// TIA Portal project "ROLLINGMILLPLC" (V16) (continued)
VERSION : 0.1
// This block is AUTO GENERATED - DO NOT MODIFY this block!
// Created by Target 1500S version 0
// at 0 
// ********************************************************
//  This is generated by Target 1500S for Simulink
//  Model name:                  LQ
//  Model version:               1.16
//                
//  ODK 1500S version:           V2.5
//  Target 1500S version:        V4.0         
//  MATLAB version:              9.9 (R2020b) 29-Jul-2020
//  Simulink version:            10.2 (R2020b) 29-Jul-2020
//  MATLAB Coder version:        5.1 (R2020b) 29-Jul-2020
//  Simulink Coder version:      9.4 (R2020b) 29-Jul-2020
// 
//  ***Model details***
//  Step Size:                   0.01
//  Default parameter behaviour: Tunable 
//  External Mode:               Off
//  ***ODK 1500S details***  
//  Heap Size:                   32k
//  Max Block Size:              1024
//  Size of thread stack:        32k
//  SyncCallParallelCount:       1(max. number of parallel calls into this ODK application)
//  ********************************************************
// Call this FB to establish a connection to user defined Web page.
   VAR_INPUT
      InternalSignals : "LQInternalModelSignals";
      CTRL_DB : DB_WWW;
   END_VAR
   VAR_IN_OUT
      Params : "LQParams";
   END_VAR
   VAR
      TestPointedSignals : "LQInternalModelSignals";
      Parameter : "LQParams";
      RWParams_Instance : "LQReadWriteParameters";
      Write : Int := 0;
      RunTime : LReal;
   END_VAR
   VAR_TEMP
      ret : Int;
   END_VAR
BEGIN
   // This is generated by Target 1500S for Simulink
   // Model name:                  LQ
   // Model version:               1.16
   //               
   // ODK 1500S version:           V2.5
   // Target 1500S version:        V4.0         
   // MATLAB version:              9.9 (R2020b) 29-Jul-2020
   // Simulink version:            10.2 (R2020b) 29-Jul-2020
   // MATLAB Coder version:        5.1 (R2020b) 29-Jul-2020
   // Simulink Coder version:      9.4 (R2020b) 29-Jul-2020
   //
   // ***Model details***
   // Step Size:                   0.01
   // Default parameter behaviour: Tunable 
   // External Mode:               Off
   // ***ODK 1500S details***  
   // Heap Size:                   32k
   // Max Block Size:              1024
   // Size of thread stack:        32k
   // SyncCallParallelCount:       1(max. number of parallel calls into this ODK application)
   // ********************************************************
   //Call this FB to establish a connection to user defined Web page.
   #RunTime := #RunTime + 10.0;

   #TestPointedSignals := #InternalSignals;
   CASE #Write OF
       0:
           #RWParams_Instance(write := FALSE,
                              STATUS => #RWParams_Instance.STATUS,
                              inOutParams := #Parameter);
           #Params := #Parameter;
       1:
           // Wait for parameter be updated by the Web action
           ;
       2:
           #RWParams_Instance(write := TRUE,
                              STATUS => #RWParams_Instance.STATUS,
                              inOutParams := #Parameter);
           #Params := #Parameter;
           #Write := 0;
       ELSE
           // Not possible to reach
           ;
   END_CASE;

   #ret := WWW(#CTRL_DB);
END_FUNCTION_BLOCK

ORGANIZATION_BLOCK "Main"   // OB1, LAD, ProgramCycle
TITLE = "Main Program Sweep (Cycle)"
{ S7_Optimized_Access := 'TRUE' }
VERSION : 0.1
   VAR_INPUT
      Initial_Call : Bool;   // Initial call of this OB
      Remanence : Bool;   // =True, if remanent data are available
   END_VAR
BEGIN
END_ORGANIZATION_BLOCK

ORGANIZATION_BLOCK "Cyclic interrupt"   // OB30, LAD, CyclicInterrupt
{ S7_Optimized_Access := 'TRUE' }
VERSION : 0.1
   VAR_INPUT
      Initial_Call : Bool;   // Initial call of this OB
      Event_Count : Int;   // Events discarded
   END_VAR
BEGIN

REGION Network 1 (SCL)
   "LQ_GlobalData".Feedback := "OpcInterface".Feedback;
END_REGION

REGION Network 2
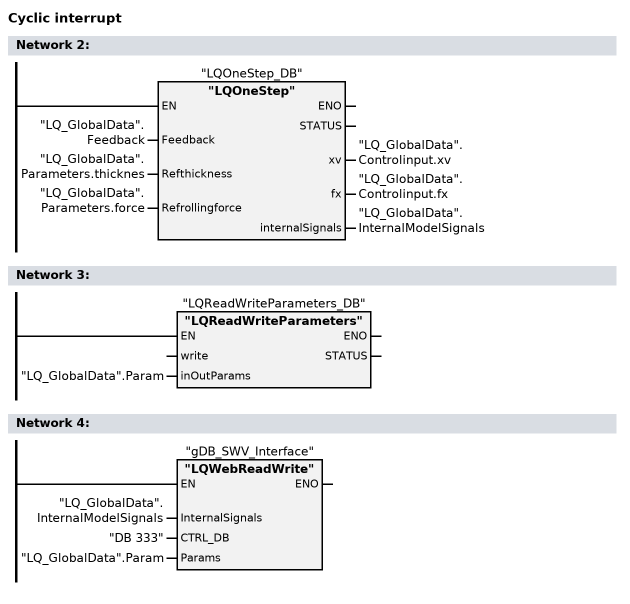
   RUNG wire#powerrail
      "LQOneStep_DB"(Feedback := "LQ_GlobalData".Feedback, Refthickness := "LQ_GlobalData".Parameters.thicknes, Refrollingforce := "LQ_GlobalData".Parameters.force, STATUS =>, xv => "LQ_GlobalData".Controlinput.xv, fx => "LQ_GlobalData".Controlinput.fx, internalSignals => "LQ_GlobalData".InternalModelSignals)
   END_RUNG
   // the same network as SCL:
   "LQOneStep_DB"(Feedback := "LQ_GlobalData".Feedback,   // "LQOneStep"
                  Refthickness := "LQ_GlobalData".Parameters.thicknes,
                  Refrollingforce := "LQ_GlobalData".Parameters.force,
                  xv => "LQ_GlobalData".Controlinput.xv,
                  fx => "LQ_GlobalData".Controlinput.fx,
                  internalSignals => "LQ_GlobalData".InternalModelSignals);
END_REGION

REGION Network 3
   RUNG wire#powerrail
      "LQReadWriteParameters_DB"(write :=, inOutParams := "LQ_GlobalData".Param, STATUS =>)
   END_RUNG
   // the same network as SCL:
   "LQReadWriteParameters_DB"(inOutParams := "LQ_GlobalData".Param);   // "LQReadWriteParameters"
END_REGION

REGION Network 4
   RUNG wire#powerrail
      "gDB_SWV_Interface"(InternalSignals := "LQ_GlobalData".InternalModelSignals, CTRL_DB := "DB 333", Params := "LQ_GlobalData".Param)
   END_RUNG
   // the same network as SCL:
   "gDB_SWV_Interface"(InternalSignals := "LQ_GlobalData".InternalModelSignals,   // "LQWebReadWrite"
                       CTRL_DB := "DB 333",
                       Params := "LQ_GlobalData".Param);
END_REGION

REGION Network 5 (SCL)
   "OpcInterface".Controlinput.xv := "LQ_GlobalData".Controlinput.xv;
   "OpcInterface".Controlinput.fx := "LQ_GlobalData".Controlinput.fx;
END_REGION
END_ORGANIZATION_BLOCK

ORGANIZATION_BLOCK "Startup"   // OB100, LAD, Startup
TITLE = "Complete Restart"
{ S7_Optimized_Access := 'TRUE' }
VERSION : 0.1
   VAR_INPUT
      LostRetentive : Bool;   // True if retentive data are lost
      LostRTC : Bool;   // True if date and time are lost
   END_VAR
BEGIN

REGION Network 1
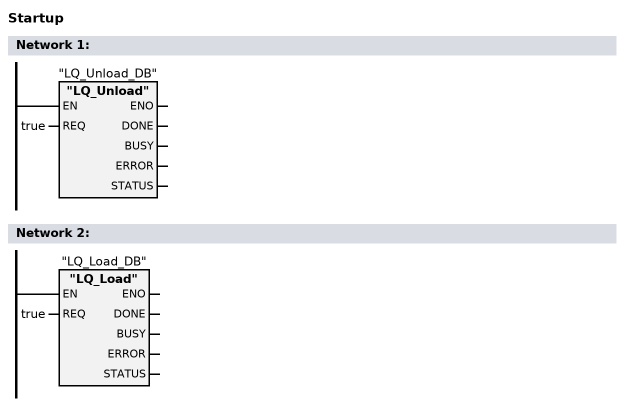
   RUNG wire#powerrail
      "LQ_Unload_DB"(REQ := true, DONE =>, BUSY =>, ERROR =>, STATUS =>)
   END_RUNG
   // the same network as SCL:
   "LQ_Unload_DB"(REQ := true);   // "LQ_Unload"
END_REGION

REGION Network 2
   RUNG wire#powerrail
      "LQ_Load_DB"(REQ := true, DONE =>, BUSY =>, ERROR =>, STATUS =>)
   END_RUNG
   // the same network as SCL:
   "LQ_Load_DB"(REQ := true);   // "LQ_Load"
END_REGION
END_ORGANIZATION_BLOCK

// ===== PLC "PLC_3"  CPU 1518-4 PN/DP MFP =====

TYPE "LQInternalModelSignals"
// This block is AUTO GENERATED - DO NOT MODIFY this block!
// Created by ODK_CodeGenerator version 205.100.101.18
// at Fri August 27 01:33:44 2021
// ********************************************************
   STRUCT
      Controlinput : Array[0..1] of LReal;
      Feedback : Array[0..4] of LReal;
      LQ_Refthickness : LReal;
      LQ_Refrollingforce : LReal;
   END_STRUCT;
END_TYPE

TYPE "LQParams"
// This block is AUTO GENERATED - DO NOT MODIFY this block!
// Created by ODK_CodeGenerator version 205.100.101.18
// at Mon August 30 17:02:50 2021
// ********************************************************
   STRUCT
      Lr : Array[0..3] of LReal;   // [LQ Controller 1/Gain Lr]:LQ_P.Lr
      Ly : Array[0..9] of LReal;   // [LQ Controller 1/Gain Ly]:LQ_P.Ly
   END_STRUCT;
   // Lr[0] := 0.013106;
   // Lr[1] := 0.0;
   // Lr[2] := 0.0;
   // Lr[3] := 3.112673;
   // Ly[0] := 0.0;
   // Ly[1] := 0.0;
   // Ly[2] := 0.0;
   // Ly[3] := 0.0;
   // Ly[4] := 0.011684;
   // Ly[5] := 0.0;
   // Ly[6] := 3.8E-05;
   // Ly[7] := 0.0;
   // Ly[8] := 0.0;
   // Ly[9] := 3.112673;
END_TYPE

DATA_BLOCK "LQ_GlobalData"   // DB1
{ S7_Optimized_Access := 'TRUE' }
VERSION : 0.1
   VAR
      Parameters : Struct
         thicknes : LReal;
         force : LReal;
      END_STRUCT;
      Feedback : Array[0..4] of LReal;
      Controlinput : Struct
         xv : LReal;
         fx : LReal;
      END_STRUCT;
      InternalModelSignals : "LQInternalModelSignals";
   END_VAR
   VAR RETAIN
      Param : "LQParams";
   END_VAR
BEGIN
END_DATA_BLOCK

DATA_BLOCK "gDB_SWV_Interface"   // DB2
{ S7_Optimized_Access := 'TRUE' }
VERSION : 0.1
// stored: InstanceOfName LQWebReadWrite
"LQWebReadWrite"
BEGIN
END_DATA_BLOCK

DATA_BLOCK "OpcInterface"   // DB3
{ S7_Optimized_Access := 'TRUE' }
VERSION : 0.1
   VAR
      Feedback : Array[0..4] of LReal;
      Controlinput : Struct
         xv : LReal;
         fx : LReal;
      END_STRUCT;
   END_VAR
BEGIN
END_DATA_BLOCK

DATA_BLOCK "LQ_Load_DB"   // DB4
{ S7_Optimized_Access := 'TRUE' }
VERSION : 0.1
// stored: InstanceOfName LQ_Load
"LQ_Load"
BEGIN
END_DATA_BLOCK

DATA_BLOCK "LQOneStep_DB"   // DB5
{ S7_Optimized_Access := 'TRUE' }
VERSION : 0.1
// stored: InstanceOfName LQOneStep
"LQOneStep"
BEGIN
END_DATA_BLOCK

DATA_BLOCK "LQReadWriteParameters_DB"   // DB6
{ S7_Optimized_Access := 'TRUE' }
VERSION : 0.1
// stored: InstanceOfName LQReadWriteParameters
"LQReadWriteParameters"
BEGIN
END_DATA_BLOCK

DATA_BLOCK "LQ_Unload_DB"   // DB7
{ S7_Optimized_Access := 'TRUE' }
VERSION : 0.1
// stored: InstanceOfName LQ_Unload
"LQ_Unload"
BEGIN
END_DATA_BLOCK

FUNCTION_BLOCK "LQ_Load"   // FB1, SCL
{ S7_Optimized_Access := 'TRUE' }
VERSION : 0.1
// This block is AUTO GENERATED - DO NOT MODIFY this block!
// Created by ODK_CodeGenerator version 2.5.1
// at Fri August 27 01:33:44 2021
// max. number of parallel calls into this ODK application is: 1
// *************************************************************
   VAR_INPUT
      REQ : Bool;
   END_VAR
   VAR_OUTPUT
      DONE : Bool;
      BUSY : Bool;
      ERROR : Bool;
      STATUS : Int;
   END_VAR
   VAR
      ODK_Load_Instance : ODK_Load;
      _odk_internal_LIBRARY_NAME : String := '<rt>LQ_ODK.so';
   END_VAR
   VAR CONSTANT
      _odk_internal_INSTANCE_ID : UDInt := 101_277_234;
   END_VAR
BEGIN
   //
   // DO NOT CHANGE BELOW OF THIS LINE !!
   // This is an automatic generated block by the
   // SIMATIC ODK 1500S V2.5.1
   // DO NOT CHANGE !!
   //
   #ODK_Load_Instance(REQ := #REQ,
                      LIBRARY_NAME := #_odk_internal_LIBRARY_NAME,
                      INSTANCE_ID := #_odk_internal_INSTANCE_ID,
                      DONE => #DONE,
                      BUSY => #BUSY,
                      ERROR => #ERROR,
                      STATUS => #STATUS);
   //
   // DO NOT CHANGE !!
   // This is an automatic generated block by the
   // SIMATIC ODK 1500S V2.5.1
   // DO NOT CHANGE ABOVE OF THIS LINE !!
   //
END_FUNCTION_BLOCK

FUNCTION_BLOCK "LQ_Unload"   // FB2, SCL
{ S7_Optimized_Access := 'TRUE' }
VERSION : 0.1
// This block is AUTO GENERATED - DO NOT MODIFY this block!
// Created by ODK_CodeGenerator version 205.100.101.18
// at Fri August 27 01:33:44 2021
// max. number of parallel calls into this ODK application is: 1
// *************************************************************
   VAR_INPUT
      REQ : Bool;
   END_VAR
   VAR_OUTPUT
      DONE : Bool;
      BUSY : Bool;
      ERROR : Bool;
      STATUS : Int;
   END_VAR
   VAR
      ODK_Unld_Instance : ODK_Unld;
   END_VAR
   VAR CONSTANT
      _odk_internal_INSTANCE_ID : UDInt := 101_277_234;
   END_VAR
BEGIN
   //
   // DO NOT CHANGE BELOW OF THIS LINE !!
   // This is an automatic generated block by the
   // SIMATIC ODK 1500S V2.5.1
   // DO NOT CHANGE !!
   //
   #ODK_Unld_Instance(REQ := #REQ,
                      INSTANCE_ID := #_odk_internal_INSTANCE_ID,
                      DONE => #DONE,
                      BUSY => #BUSY,
                      ERROR => #ERROR,
                      STATUS => #STATUS);
   //
   // DO NOT CHANGE !!
   // This is an automatic generated block by the
   // SIMATIC ODK 1500S V2.5.1
   // DO NOT CHANGE ABOVE OF THIS LINE !!
   //
END_FUNCTION_BLOCK

FUNCTION_BLOCK "LQOneStep"   // FB3, SCL
{ S7_Optimized_Access := 'TRUE' }
VERSION : 0.1
// This block is AUTO GENERATED - DO NOT MODIFY this block!
// Created by ODK_CodeGenerator version 205.100.101.18
// at Fri August 27 01:33:44 2021
// max. number of parallel calls into this ODK application is: 1
// *************************************************************
//  This is generated by Target 1500S for Simulink
//  Model name:                  LQ
//  Model version:               1.16
//                 
//  ODK 1500S version:           V2.5
//  Target 1500S version:        V4.0         
//  MATLAB version:              9.9 (R2020b) 29-Jul-2020
//  Simulink version:            10.2 (R2020b) 29-Jul-2020
//  MATLAB Coder version:        5.1 (R2020b) 29-Jul-2020
//  Simulink Coder version:      9.4 (R2020b) 29-Jul-2020
//  
//  ***Model details***
//  Step Size:                   0.01
//  Default parameter behaviour: Tunable
//  External Mode:               Off
//  
//  ***ODK 1500S details***  
//  Heap Size:                   32k
//  Max Block Size:              1024
//  Size of thread stack:        32k
//  SyncCallParallelCount:       1(max. number of parallel calls into this ODK application)
//  ********************************************************
   VAR_INPUT
      Feedback : Array[0..4] of LReal;
      Refthickness : LReal;
      Refrollingforce : LReal;
   END_VAR
   VAR_OUTPUT
      STATUS : Int := 0;
      xv : LReal;
      fx : LReal;
      internalSignals : "LQInternalModelSignals";
   END_VAR
   VAR
      _odk_internal_Last_REQ : Bool := FALSE;
      _odk_internal_Last_BUSY : Bool := FALSE;
      _odk_internal_IN_BUFFER : Array[0..55] of Byte;
      _odk_internal_OUT_BUFFER : Array[0..87] of Byte;
   END_VAR
   VAR_TEMP
      _odk_internal_pos : DInt;
      _odk_internal_err : Int;
      _odk_internal_i : Int;
   END_VAR
   VAR CONSTANT
      _odk_internal_INSTANCE_ID : UDInt := 101_277_234;
      _odk_internal_COMMAND : UDInt := 295_977_560;
   END_VAR
BEGIN
   //
   // DO NOT CHANGE BELOW OF THIS LINE !!
   // This is an automatic generated block by the
   // SIMATIC ODK 1500S V2.5.1
   // DO NOT CHANGE !!
   //
   // This is generated by Target 1500S for Simulink
   // Model name:                  LQ
   // Model version:               1.16
   //                
   // ODK 1500S version:           V2.5
   // Target 1500S version:        V4.0         
   // MATLAB version:              9.9 (R2020b) 29-Jul-2020
   // Simulink version:            10.2 (R2020b) 29-Jul-2020
   // MATLAB Coder version:        5.1 (R2020b) 29-Jul-2020
   // Simulink Coder version:      9.4 (R2020b) 29-Jul-2020
   // 
   // ***Model details***
   // Step Size:                   0.01
   // Default parameter behaviour: Tunable
   // External Mode:               Off
   // 
   // ***ODK 1500S details***  
   // Heap Size:                   32k
   // Max Block Size:              1024
   // Size of thread stack:        32k
   // SyncCallParallelCount:       1(max. number of parallel calls into this ODK application)
   // ********************************************************
   // 
   #_odk_internal_pos := 0;
   FOR #_odk_internal_i := 0 TO 4 DO
       #_odk_internal_err := WRITE_LITTLE(src_variable := #Feedback[#_odk_internal_i], dest_array := #_odk_internal_IN_BUFFER, pos := #_odk_internal_pos);
   END_FOR;
   #_odk_internal_err := WRITE_LITTLE(src_variable := #Refthickness, dest_array := #_odk_internal_IN_BUFFER, pos := #_odk_internal_pos);
   #_odk_internal_err := WRITE_LITTLE(src_variable := #Refrollingforce, dest_array := #_odk_internal_IN_BUFFER, pos := #_odk_internal_pos);
   #STATUS := ODK_ExcS(INSTANCE_ID := #_odk_internal_INSTANCE_ID,
                       COMMAND := #_odk_internal_COMMAND,
                       IN_DATA := #_odk_internal_IN_BUFFER,
                       INOUT_DATA := null,
                       OUT_DATA := #_odk_internal_OUT_BUFFER
   );
   IF INT_TO_UINT(#STATUS) < 16#7000 THEN
       #_odk_internal_pos := 0;
       #_odk_internal_err := READ_LITTLE(dest_Variable => #xv, src_array := #_odk_internal_OUT_BUFFER, pos := #_odk_internal_pos);
       #_odk_internal_err := READ_LITTLE(dest_Variable => #fx, src_array := #_odk_internal_OUT_BUFFER, pos := #_odk_internal_pos);
       FOR #_odk_internal_i := 0 TO 1 DO
           #_odk_internal_err := READ_LITTLE(dest_Variable => #internalSignals.#Controlinput[#_odk_internal_i], src_array := #_odk_internal_OUT_BUFFER, pos := #_odk_internal_pos);
       END_FOR;
       FOR #_odk_internal_i := 0 TO 4 DO
           #_odk_internal_err := READ_LITTLE(dest_Variable => #internalSignals.#Feedback[#_odk_internal_i], src_array := #_odk_internal_OUT_BUFFER, pos := #_odk_internal_pos);
       END_FOR;
       #_odk_internal_err := READ_LITTLE(dest_Variable => #internalSignals.#LQ_Refthickness, src_array := #_odk_internal_OUT_BUFFER, pos := #_odk_internal_pos);
       #_odk_internal_err := READ_LITTLE(dest_Variable => #internalSignals.#LQ_Refrollingforce, src_array := #_odk_internal_OUT_BUFFER, pos := #_odk_internal_pos);
   END_IF;
   //
   // DO NOT CHANGE !!
   // This is an automatic generated block by the
   // SIMATIC ODK 1500S V2.5.1
   // DO NOT CHANGE ABOVE OF THIS LINE !!
   //
END_FUNCTION_BLOCK

FUNCTION_BLOCK "LQReadWriteParameters"   // FB4, SCL
{ S7_Optimized_Access := 'TRUE' }
VERSION : 0.1
// This block is AUTO GENERATED - DO NOT MODIFY this block!
// Created by ODK_CodeGenerator version 205.100.101.18
// at Fri August 27 01:33:44 2021
// max. number of parallel calls into this ODK application is: 1
// *************************************************************
//  This is generated by Target 1500S for Simulink
//  Model name:                  LQ
//  Model version:               1.16
//                 
//  ODK 1500S version:           V2.5
//  Target 1500S version:        V4.0         
//  MATLAB version:              9.9 (R2020b) 29-Jul-2020
//  Simulink version:            10.2 (R2020b) 29-Jul-2020
//  MATLAB Coder version:        5.1 (R2020b) 29-Jul-2020
//  Simulink Coder version:      9.4 (R2020b) 29-Jul-2020
//  
//  ***Model details***
//  Step Size:                   0.01
//  Default parameter behaviour: Tunable
//  External Mode:               Off
//  
//  ***ODK 1500S details***  
//  Heap Size:                   32k
//  Max Block Size:              1024
//  Size of thread stack:        32k
//  SyncCallParallelCount:       1(max. number of parallel calls into this ODK application)
//  ********************************************************
//  
//  Call this function to read or write parameters from/to Simulink Model.
//  Set write[IN] parameter to TRUE in order to write and set FALSE to read parameters
   VAR_INPUT
      write : Bool;
   END_VAR
   VAR_OUTPUT
      STATUS : Int := 0;
   END_VAR
   VAR_IN_OUT
      inOutParams : "LQParams";
   END_VAR
   VAR
      _odk_internal_Last_REQ : Bool := FALSE;
      _odk_internal_Last_BUSY : Bool := FALSE;
      _odk_internal_IN_BUFFER : Array[0..0] of Byte;
      _odk_internal_INOUT_BUFFER : Array[0..111] of Byte;
   END_VAR
   VAR_TEMP
      _odk_internal_pos : DInt;
      _odk_internal_err : Int;
      _odk_internal_i : Int;
   END_VAR
   VAR CONSTANT
      _odk_internal_INSTANCE_ID : UDInt := 101_277_234;
      _odk_internal_COMMAND : UDInt := 2_137_970_399;
   END_VAR
BEGIN
   //
   // DO NOT CHANGE BELOW OF THIS LINE !!
   // This is an automatic generated block by the
   // SIMATIC ODK 1500S V2.5.1
   // DO NOT CHANGE !!
   //
   // This is generated by Target 1500S for Simulink
   // Model name:                  LQ
   // Model version:               1.16
   //                
   // ODK 1500S version:           V2.5
   // Target 1500S version:        V4.0         
   // MATLAB version:              9.9 (R2020b) 29-Jul-2020
   // Simulink version:            10.2 (R2020b) 29-Jul-2020
   // MATLAB Coder version:        5.1 (R2020b) 29-Jul-2020
   // Simulink Coder version:      9.4 (R2020b) 29-Jul-2020
   // 
   // ***Model details***
   // Step Size:                   0.01
   // Default parameter behaviour: Tunable
   // External Mode:               Off
   // 
   // ***ODK 1500S details***  
   // Heap Size:                   32k
   // Max Block Size:              1024
   // Size of thread stack:        32k
   // SyncCallParallelCount:       1(max. number of parallel calls into this ODK application)
   // ********************************************************
   // 
   // Call this function to read or write parameters from/to Simulink Model.
   // Set write[IN] parameter to TRUE in order to write and set FALSE to read parameters
   #_odk_internal_pos := 0;
   IF (True = #write) THEN
       #_odk_internal_IN_BUFFER[#_odk_internal_pos] := BYTE#1;
   ELSE
       #_odk_internal_IN_BUFFER[#_odk_internal_pos] := BYTE#0;
   END_IF;
   #_odk_internal_pos := #_odk_internal_pos + 1;
   #_odk_internal_pos := 0;
   FOR #_odk_internal_i := 0 TO 3 DO
       #_odk_internal_err := WRITE_LITTLE(src_variable := #inOutParams.#Lr[#_odk_internal_i], dest_array := #_odk_internal_INOUT_BUFFER, pos := #_odk_internal_pos);
   END_FOR;
   FOR #_odk_internal_i := 0 TO 9 DO
       #_odk_internal_err := WRITE_LITTLE(src_variable := #inOutParams.#Ly[#_odk_internal_i], dest_array := #_odk_internal_INOUT_BUFFER, pos := #_odk_internal_pos);
   END_FOR;
   #STATUS := ODK_ExcS(INSTANCE_ID := #_odk_internal_INSTANCE_ID,
                       COMMAND := #_odk_internal_COMMAND,
                       IN_DATA := #_odk_internal_IN_BUFFER,
                       INOUT_DATA := #_odk_internal_INOUT_BUFFER,
                       OUT_DATA := null);
   IF INT_TO_UINT(#STATUS) < 16#7000 THEN
       #_odk_internal_pos := 0;
       FOR #_odk_internal_i := 0 TO 3 DO
           #_odk_internal_err := READ_LITTLE(dest_Variable => #inOutParams.#Lr[#_odk_internal_i], src_array := #_odk_internal_INOUT_BUFFER, pos := #_odk_internal_pos);
       END_FOR;
       FOR #_odk_internal_i := 0 TO 9 DO
           #_odk_internal_err := READ_LITTLE(dest_Variable => #inOutParams.#Ly[#_odk_internal_i], src_array := #_odk_internal_INOUT_BUFFER, pos := #_odk_internal_pos);
       END_FOR;
   END_IF;
   //
   // DO NOT CHANGE !!
   // This is an automatic generated block by the
   // SIMATIC ODK 1500S V2.5.1
   // DO NOT CHANGE ABOVE OF THIS LINE !!
   //
END_FUNCTION_BLOCK

FUNCTION_BLOCK "LQWebReadWrite"   // FB5, SCL
{ S7_Optimized_Access := 'TRUE' }
VERSION : 0.1
// This block is AUTO GENERATED - DO NOT MODIFY this block!
// Created by Target 1500S version 0
// at 0 
// ********************************************************
//  This is generated by Target 1500S for Simulink
//  Model name:                  LQ
//  Model version:               1.16
//                
//  ODK 1500S version:           V2.5
//  Target 1500S version:        V4.0         
//  MATLAB version:              9.9 (R2020b) 29-Jul-2020
//  Simulink version:            10.2 (R2020b) 29-Jul-2020
//  MATLAB Coder version:        5.1 (R2020b) 29-Jul-2020
//  Simulink Coder version:      9.4 (R2020b) 29-Jul-2020
// 
//  ***Model details***
//  Step Size:                   0.01
//  Default parameter behaviour: Tunable 
//  External Mode:               Off
//  ***ODK 1500S details***  
//  Heap Size:                   32k
//  Max Block Size:              1024
//  Size of thread stack:        32k
//  SyncCallParallelCount:       1(max. number of parallel calls into this ODK application)
//  ********************************************************
// Call this FB to establish a connection to user defined Web page.
   VAR_INPUT
      InternalSignals : "LQInternalModelSignals";
      CTRL_DB : DB_WWW;
   END_VAR
   VAR_IN_OUT
      Params : "LQParams";
   END_VAR
   VAR
      TestPointedSignals : "LQInternalModelSignals";
      Parameter : "LQParams";
      RWParams_Instance : "LQReadWriteParameters";
      Write : Int := 0;
      RunTime : LReal;
   END_VAR
   VAR_TEMP
      ret : Int;
   END_VAR
BEGIN
   // This is generated by Target 1500S for Simulink
   // Model name:                  LQ
   // Model version:               1.16
   //               
   // ODK 1500S version:           V2.5
   // Target 1500S version:        V4.0         
   // MATLAB version:              9.9 (R2020b) 29-Jul-2020
   // Simulink version:            10.2 (R2020b) 29-Jul-2020
   // MATLAB Coder version:        5.1 (R2020b) 29-Jul-2020
   // Simulink Coder version:      9.4 (R2020b) 29-Jul-2020
   //
   // ***Model details***
   // Step Size:                   0.01
   // Default parameter behaviour: Tunable 
   // External Mode:               Off
   // ***ODK 1500S details***  
   // Heap Size:                   32k
   // Max Block Size:              1024
   // Size of thread stack:        32k
   // SyncCallParallelCount:       1(max. number of parallel calls into this ODK application)
   // ********************************************************
   //Call this FB to establish a connection to user defined Web page.
   #RunTime := #RunTime + 10.0;

   #TestPointedSignals := #InternalSignals;
   CASE #Write OF
       0:
           #RWParams_Instance(write := FALSE,
                              STATUS => #RWParams_Instance.STATUS,
                              inOutParams := #Parameter);
           #Params := #Parameter;
       1:
           // Wait for parameter be updated by the Web action
           ;
       2:
           #RWParams_Instance(write := TRUE,
                              STATUS => #RWParams_Instance.STATUS,
                              inOutParams := #Parameter);
           #Params := #Parameter;
           #Write := 0;
       ELSE
           // Not possible to reach
           ;
   END_CASE;

   #ret := WWW(#CTRL_DB);
END_FUNCTION_BLOCK

ORGANIZATION_BLOCK "Main"   // OB1, LAD, ProgramCycle
TITLE = "Main Program Sweep (Cycle)"
{ S7_Optimized_Access := 'TRUE' }
VERSION : 0.1
   VAR_INPUT
      Initial_Call : Bool;   // Initial call of this OB
      Remanence : Bool;   // =True, if remanent data are available
   END_VAR
BEGIN
END_ORGANIZATION_BLOCK

ORGANIZATION_BLOCK "Cyclic interrupt"   // OB30, LAD, CyclicInterrupt
{ S7_Optimized_Access := 'TRUE' }
VERSION : 0.1
   VAR_INPUT
      Initial_Call : Bool;   // Initial call of this OB
      Event_Count : Int;   // Events discarded
   END_VAR
BEGIN

REGION Network 1 (SCL)
   "LQ_GlobalData".Feedback := "OpcInterface".Feedback;
END_REGION

REGION Network 2
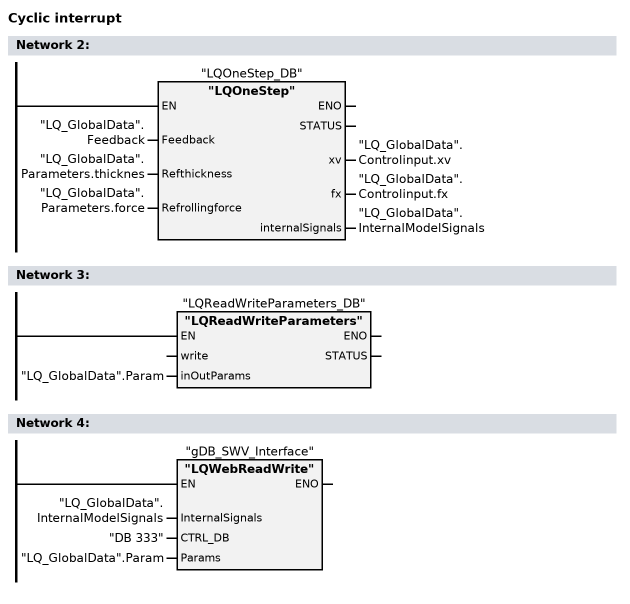
   RUNG wire#powerrail
      "LQOneStep_DB"(Feedback := "LQ_GlobalData".Feedback, Refthickness := "LQ_GlobalData".Parameters.thicknes, Refrollingforce := "LQ_GlobalData".Parameters.force, STATUS =>, xv => "LQ_GlobalData".Controlinput.xv, fx => "LQ_GlobalData".Controlinput.fx, internalSignals => "LQ_GlobalData".InternalModelSignals)
   END_RUNG
   // the same network as SCL:
   "LQOneStep_DB"(Feedback := "LQ_GlobalData".Feedback,   // "LQOneStep"
                  Refthickness := "LQ_GlobalData".Parameters.thicknes,
                  Refrollingforce := "LQ_GlobalData".Parameters.force,
                  xv => "LQ_GlobalData".Controlinput.xv,
                  fx => "LQ_GlobalData".Controlinput.fx,
                  internalSignals => "LQ_GlobalData".InternalModelSignals);
END_REGION

REGION Network 3
   RUNG wire#powerrail
      "LQReadWriteParameters_DB"(write :=, inOutParams := "LQ_GlobalData".Param, STATUS =>)
   END_RUNG
   // the same network as SCL:
   "LQReadWriteParameters_DB"(inOutParams := "LQ_GlobalData".Param);   // "LQReadWriteParameters"
END_REGION

REGION Network 4
   RUNG wire#powerrail
      "gDB_SWV_Interface"(InternalSignals := "LQ_GlobalData".InternalModelSignals, CTRL_DB := "DB 333", Params := "LQ_GlobalData".Param)
   END_RUNG
   // the same network as SCL:
   "gDB_SWV_Interface"(InternalSignals := "LQ_GlobalData".InternalModelSignals,   // "LQWebReadWrite"
                       CTRL_DB := "DB 333",
                       Params := "LQ_GlobalData".Param);
END_REGION

REGION Network 5 (SCL)
   "OpcInterface".Controlinput.xv := "LQ_GlobalData".Controlinput.xv;
   "OpcInterface".Controlinput.fx := "LQ_GlobalData".Controlinput.fx;
END_REGION
END_ORGANIZATION_BLOCK

ORGANIZATION_BLOCK "Startup"   // OB100, LAD, Startup
TITLE = "Complete Restart"
{ S7_Optimized_Access := 'TRUE' }
VERSION : 0.1
   VAR_INPUT
      LostRetentive : Bool;   // True if retentive data are lost
      LostRTC : Bool;   // True if date and time are lost
   END_VAR
BEGIN

REGION Network 1
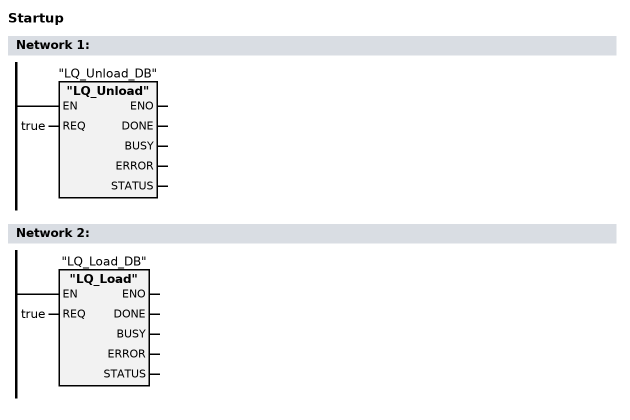
   RUNG wire#powerrail
      "LQ_Unload_DB"(REQ := true, DONE =>, BUSY =>, ERROR =>, STATUS =>)
   END_RUNG
   // the same network as SCL:
   "LQ_Unload_DB"(REQ := true);   // "LQ_Unload"
END_REGION

REGION Network 2
   RUNG wire#powerrail
      "LQ_Load_DB"(REQ := true, DONE =>, BUSY =>, ERROR =>, STATUS =>)
   END_RUNG
   // the same network as SCL:
   "LQ_Load_DB"(REQ := true);   // "LQ_Load"
END_REGION
END_ORGANIZATION_BLOCK

(* ===== HMI "HMI_RT_2" =====
system functions are stored by id; their names below are inferred from use
connection "HMI_Connection_1": ETHERNET, S7_1500_OMS
connection "HMI_Connection_2": ETHERNET, S7_1500_OMS
connection "HMI_Connection_3": ETHERNET, S7_1500_OMS

HMI tags "Default tag table"
   "Tag_ScreenNumber" : UInt, internal
   "LQ_GlobalData_Parameters_thicknes" : LReal = PLC LQ_GlobalData.Parameters.thicknes, 1 s
   "LQ_GlobalData_Parameters_force" : LReal = PLC LQ_GlobalData.Parameters.force, 1 s
   "LQ_GlobalData_Feedback{2}" : LReal = PLC LQ_GlobalData.Feedback[2], 1 s
   "LQ_GlobalData_Parameters_thicknes(1)" : LReal = PLC LQ_GlobalData.Parameters.thicknes, 1 s
   "LQ_GlobalData_Feedback{2}(1)" : LReal = PLC LQ_GlobalData.Feedback[2], 1 s
   "LQ_GlobalData_Parameters_force(1)" : LReal = PLC LQ_GlobalData.Parameters.force, 1 s
   "LQ_GlobalData_Parameters_thicknes(2)" : LReal = PLC LQ_GlobalData.Parameters.thicknes, 1 s
   "LQ_GlobalData_Parameters_force(2)" : LReal = PLC LQ_GlobalData.Parameters.force, 1 s
   "LQ_GlobalData_Feedback{2}(2)" : LReal = PLC LQ_GlobalData.Feedback[2], 1 s
   "LQ_GlobalData_Feedback{4}" : LReal = PLC LQ_GlobalData.Feedback[4], 1 s
   "LQ_GlobalData_Feedback{4}(1)" : LReal = PLC LQ_GlobalData.Feedback[4], 1 s
   "LQ_GlobalData_Feedback{4}(2)" : LReal = PLC LQ_GlobalData.Feedback[4], 1 s

screen "Home" 1280x740, template "Template_1"
   on GenerateScreen: SetTag("Tag_ScreenNumber", 1)
   TextField "HmiScreenItemData_3" at 413,45 size 404x37; Text 'Welcome to HMI of the Rolling Mill'
   Button "HmiScreenItemData" at 471,181 size 159x47; TextOn 'Rolling Stand 1'; TextOff 'Rolling Stand 1'; PictureOn "Navigates to Roller 1 for TP1500 Comfort 16.0.0.0"; PictureOff "Navigates to Roller 1 for TP1500 Comfort 16.0.0.0"
      on Release: ActivateScreen("Rolling Stand 1", 0)
   Button "HmiScreenItemData_1" at 471,261 size 159x47; TextOn 'Rolling Stand 2'; TextOff 'Rolling Stand 2'; PictureOn "Navigates to Roller 2 for TP1500 Comfort 16.0.0.0"; PictureOff "Navigates to Roller 2 for TP1500 Comfort 16.0.0.0"
      on Release: ActivateScreen("Rolling Stand 2", 0)
   Button "HmiScreenItemData_2" at 471,342 size 159x47; TextOn 'Rolling Stand 3'; TextOff 'Rolling Stand 3'; PictureOn "Navigates to Roller 3 for TP1500 Comfort 16.0.0.0"; PictureOff "Navigates to Roller 3 for TP1500 Comfort 16.0.0.0"
      on Release: ActivateScreen("Rolling Stand 3", 0)
   Button "HmiScreenItemData_4" at 538,476 size 159x47; TextOn 'System screens'; TextOff 'System screens'; PictureOn "Navigates to System screens for TP1500 Comfort 16.0.0.0"; PictureOff "Navigates to System screens for TP1500 Comfort 16.0.0.0"
      on Release: ActivateScreen("System screens", 0)
   TextField "Text field_1" at 482,193 size 30x18; Text 'R-1'
   TextField "Text field_2" at 482,275 size 30x18; Text 'R-2'
   TextField "Text field_3" at 482,356 size 30x18; Text 'R-3'
   TextField "Text field_5" at 553,432 size 135x25; Text 'Information'
   Switch "Switch_1" at 683,171 size 77x50; CaptionText 'Switch'; TextOff 'OFF'; TextOn 'ON'
      on SwitchOn: function_f249594b("HMI_Connection_1", 8)
      on SwitchOff: function_f249594b("HMI_Connection_1", 4)
   Switch "Switch_2" at 683,255 size 77x50; TextOn 'ON'; CaptionText 'Switch'; TextOff 'OFF'
      on SwitchOn: function_f249594b("HMI_Connection_2", 8)
      on SwitchOff: function_f249594b("HMI_Connection_2", 4)
   Switch "Switch_3" at 683,335 size 77x50; TextOn 'ON'; CaptionText 'Switch'; TextOff 'OFF'
      on SwitchOn: function_f249594b("HMI_Connection_3", 8)
      on SwitchOff: function_f249594b("HMI_Connection_3", 4)
   TextField "Text field_4" at 480,132 size 110x25; Text 'Mill Stands'
   TextField "Text field_6" at 675,132 size 92x25; Text 'PLC Switch'

screen "Rolling Stand 1" 1280x740, template "Template_1"
   on GenerateScreen: SetTag("Tag_ScreenNumber", 2)
   TextField "HmiScreenItemData" at 146,334 size 1024x27; Text 'Roller 1'
   Button "Back" at 1,25 size 159x47; TextOn 'Back'; TextOff 'Back'
      on Release: ActivateScreen("Home", 0)
   TrendView "Trend view_1" at 295,23 size 984x343
   TextField "Text field_4" at 41,188 size 164x40; Text 'Enter Setpoint'
   Group "Group" at 29,242 size 182x37; FormatPattern 9
   Group "Group_1" at 26,92 size 196x56
   IOField "I/O field_2" at 162,288 size 71x37; FormatPattern 999; Unit N
      ProcessValue <- "LQ_GlobalData_Parameters_force"
   TextField "Text field_3" at 25,288 size 137x37; Text 'Rolling force :'
   TrendView "Trend view_2" at 296,361 size 984x320
   IOField "I/O field_1" at 150,242 size 61x37; FormatPattern 9; Unit mm
      ProcessValue <- "LQ_GlobalData_Parameters_thicknes"
   TextField "Text field_1" at 29,242 size 121x37; Text 'Thickness :'
   TextField "Text field_2" at 26,94 size 196x53; Text 'Rolling Stand 1'

screen "System screens" 1280x740, template "Template_1"
   on GenerateScreen: SetTag("Tag_ScreenNumber", 5)
   Button "Back" at 1,25 size 159x47; TextOn 'Back'; TextOff 'Back'
      on Release: ActivateScreen("Home", 0)
   Button "HmiScreenItemData" at 36,119 size 159x47; TextOn 'SIMATIC PLC system diagnos...'; TextOff 'SIMATIC PLC system diagnos...'; PictureOn "Navigates to SIMATIC PLC system diagnostics for TP1500 Comfort 16.0.0.0"; PictureOff "Navigates to SIMATIC PLC system diagnostics for TP1500 Comfort 16.0.0.0"
      on Release: ActivateScreen("SIMATIC PLC system diagnostics", 0)
   Button "HmiScreenItemData_1" at 36,178 size 159x47; TextOn 'Project information'; TextOff 'Project information'; PictureOn "Navigates to Project information for TP1500 Comfort 16.0.0.0"; PictureOff "Navigates to Project information for TP1500 Comfort 16.0.0.0"
      on Release: ActivateScreen("Project information", 0)
   Button "HmiScreenItemData_2" at 36,237 size 159x47; TextOn 'System settings'; TextOff 'System settings'; PictureOn "Navigates to System settings for TP1500 Comfort 16.0.0.0"; PictureOff "Navigates to System settings for TP1500 Comfort 16.0.0.0"
      on Release: ActivateScreen("System settings", 0)
   Button "HmiScreenItemData_3" at 36,296 size 159x47; TextOn 'User administration'; TextOff 'User administration'; PictureOn "Navigates to User administration for TP1500 Comfort 16.0.0.0"; PictureOff "Navigates to User administration for TP1500 Comfort 16.0.0.0"
      on Release: ActivateScreen("User administration", 0)
   Button "HmiScreenItemData_4" at 36,355 size 159x47; TextOn 'System information'; TextOff 'System information'; PictureOn "Navigates to System information for TP1500 Comfort 16.0.0.0"; PictureOff "Navigates to System information for TP1500 Comfort 16.0.0.0"
      on Release: ActivateScreen("System information", 0)
   Button "HmiScreenItemData_5" at 36,414 size 159x47; TextOn 'Different jobs'; TextOff 'Different jobs'; PictureOn "Navigates to Different jobs for TP1500 Comfort 16.0.0.0"; PictureOff "Navigates to Different jobs for TP1500 Comfort 16.0.0.0"
      on Release: ActivateScreen("Different jobs", 0)

screen "SIMATIC PLC system diagnostics" 1280x740, template "Template_1"
   on GenerateScreen: SetTag("Tag_ScreenNumber", 6)
   SysDiagControl "HmiScreenItemData" at 1,73 size 1276x599
   Button "Back" at 1,25 size 159x47; TextOn 'Back'; TextOff 'Back'
      on Release: ActivateScreen("System screens", 0)

screen "Project information" 1280x740, template "Template_1"
   on GenerateScreen: SetTag("Tag_ScreenNumber", 7)
   TextField "HmiScreenItemData" at 35,75 size 171x28; Text 'Project name:'
   TextField "HmiScreenItemData_1" at 241,75 size 1004x28; Text 'Rolling_Mill_With_Three_Rollers'
   TextField "HmiScreenItemData_2" at 35,105 size 171x28; Text 'Created on:'
   TextField "HmiScreenItemData_3" at 241,105 size 1004x28; Text '5/28/2021 9:23:35 PM'
   TextField "HmiScreenItemData_4" at 35,135 size 171x28; Text 'Author:'
   TextField "HmiScreenItemData_5" at 241,135 size 1004x28; Text 'Mehrab'
   TextField "HmiScreenItemData_6" at 35,165 size 171x28; Text 'Description:'
   TextField "HmiScreenItemData_7" at 241,165 size 1004x28; Text '(not configured)'
   Button "Back" at 1,25 size 159x47; TextOn 'Back'; TextOff 'Back'
      on Release: ActivateScreen("System screens", 0)

screen "System settings" 1280x740, template "Template_1"
   on GenerateScreen: SetTag("Tag_ScreenNumber", 8)
   Button "Calibrate screen" at 36,119 size 159x47; TextOn 'Calibrate screen'; TextOff 'Calibrate screen'
      on Release: function_bc3e350c()
   Button "Clean screen" at 36,178 size 159x47; TextOn 'Clean screen'; TextOff 'Clean screen'
      on Release: function_be740847(30)
   Button "Back" at 1,25 size 159x47; TextOn 'Back'; TextOff 'Back'
      on Release: ActivateScreen("System screens", 0)

screen "User administration" 1280x740, template "Template_1"
   on GenerateScreen: SetTag("Tag_ScreenNumber", 9)
   UserView "HmiScreenItemData" at 1,73 size 1276x599
   Button "Back" at 1,25 size 159x47; TextOn 'Back'; TextOff 'Back'
      on Release: ActivateScreen("System screens", 0)

screen "System information" 1280x740, template "Template_1"
   on GenerateScreen: SetTag("Tag_ScreenNumber", 10)
   TextField "HmiScreenItemData" at 35,75 size 171x28; Text 'HMI device type:'
   TextField "HmiScreenItemData_1" at 241,75 size 1004x28; Text 'TP1500 Comfort 16.0.0.0'
   TextField "HmiScreenItemData_2" at 35,105 size 171x28; Text 'Version:'
   TextField "HmiScreenItemData_3" at 35,135 size 171x28; Text 'Connection:'
   TextField "HmiScreenItemData_4" at 241,135 size 1004x28; Text '(not configured)'
   TextField "HmiScreenItemData_5" at 35,165 size 171x28; Text 'PLC:'
   TextField "HmiScreenItemData_6" at 241,165 size 1004x28; Text '<PLC>'
   Button "Display version" at 241,105 size 1004x28; TextOn 'Display version'; TextOff 'Display version'
      on Release: function_febcb963(-1)
   Button "Back" at 1,25 size 159x47; TextOn 'Back'; TextOff 'Back'
      on Release: ActivateScreen("System screens", 0)

screen "Different jobs" 1280x740, template "Template_1"
   on GenerateScreen: SetTag("Tag_ScreenNumber", 11)
   Button "Online" at 36,119 size 159x47; TextOn 'Online'; TextOff 'Online'
      on Release: function_bb44b551(0)
   Button "Offline" at 36,178 size 159x47; TextOn 'Offline'; TextOff 'Offline'
      on Release: function_bb44b551(1)
   Button "Transfer" at 36,237 size 159x47; TextOn 'Transfer'; TextOff 'Transfer'
      on Release: function_bb44b551(2)
   Button "Toggle language" at 36,296 size 159x47; TextOn 'Toggle language'; TextOff 'Toggle language'
      on Release: function_fb9197e8(-1)
   Button "Control Panel" at 36,355 size 159x47; TextOn 'Control Panel'; TextOff 'Control Panel'
      on Release: function_f34a74f3()
   Button "Stop Runtime" at 36,414 size 159x47; TextOn 'Stop Runtime'; TextOff 'Stop Runtime'
      on Release: StopRuntime(0)
   Button "Back" at 1,25 size 159x47; TextOn 'Back'; TextOff 'Back'
      on Release: ActivateScreen("System screens", 0)

screen "Rolling Stand 2" 1280x740, template "Template_1"
   on GenerateScreen: SetTag("Tag_ScreenNumber", 3)
   TextField "HmiScreenItemData" at 146,334 size 1024x27; Text 'Roller 1'
   Button "Back" at 1,25 size 159x47; TextOn 'Back'; TextOff 'Back'
      on Release: ActivateScreen("Home", 0)
   TrendView "Trend view_1" at 295,23 size 983x338
   TextField "Text field_2" at 26,94 size 196x53; Text 'Rolling Stand 2'
   Group "Group" at 29,242 size 182x37; FormatPattern 9
   IOField "I/O field_2" at 161,289 size 69x37; FormatPattern 999; Unit N
      ProcessValue <- "LQ_GlobalData_Parameters_force(1)"
   TextField "Text field_3" at 25,289 size 137x37; Text 'Rolling force :'
   TextField "Text field_4" at 41,188 size 164x40; Text 'Enter Setpoint'
   TrendView "Trend view_2" at 295,359 size 984x322
   IOField "I/O field_1" at 150,242 size 61x37; FormatPattern 9; Unit mm
      ProcessValue <- "LQ_GlobalData_Parameters_thicknes(1)"
   TextField "Text field_1" at 29,242 size 121x37; Text 'Thickness :'

screen "Rolling Stand 3" 1280x740, template "Template_1"
   on GenerateScreen: SetTag("Tag_ScreenNumber", 4)
   TextField "HmiScreenItemData" at 146,334 size 1024x27; Text 'Roller 1'
   Button "Back" at 1,25 size 159x47; TextOn 'Back'; TextOff 'Back'
      on Release: ActivateScreen("Home", 0)
   TrendView "Trend view_1" at 296,23 size 983x344
   TextField "Text field_2" at 26,94 size 196x53; Text 'Rolling Stand 3'
   Group "Group" at 29,242 size 182x37; FormatPattern 9
   Group "Group_1" at 25,286 size 204x37; FormatPattern 9
   TextField "Text field_4" at 41,188 size 164x40; Text 'Enter Setpoint'
   TrendView "Trend view_2" at 295,362 size 984x318
   IOField "I/O field_1" at 150,242 size 61x37; FormatPattern 9; Unit mm
      ProcessValue <- "LQ_GlobalData_Parameters_thicknes(2)"
   TextField "Text field_1" at 29,242 size 121x37; Text 'Thickness :'
   IOField "I/O field_2" at 161,286 size 68x37; FormatPattern 999; Unit N
      ProcessValue <- "LQ_GlobalData_Parameters_force(2)"
   TextField "Text field_3" at 25,286 size 135x37; Text 'Rolling force :'

Template "Template_1" 1280x740
   Button "Exit" at 1200,679 size 78x59; TextOn 'Exit'; TextOff 'Exit'; PictureOn "ExitRuntime_TP1500_Comfort_TR"; PictureOff "ExitRuntime_TP1500_Comfort_TR"
      on Release: StopRuntime(0)
   Button "Log on" at 1120,679 size 78x59; TextOn 'Log on'; TextOff 'Log on'; PictureOn "Login_TP1500_Comfort_TR"; PictureOff "Login_TP1500_Comfort_TR"
      on Release: function_a2a04561()
   Button "Language" at 1040,679 size 78x59; TextOn 'Language'; TextOff 'Language'; PictureOn "ToggleLanguage_TP1500_Comfort_TR"; PictureOff "ToggleLanguage_TP1500_Comfort_TR"
      on Release: function_fb9197e8(-1)
   Button "Template_Button" at 960,679 size 78x59; TextOff 'Text'
   Button "Template_Button_1" at 880,679 size 78x59; TextOff 'Text'
   Button "Template_Button_2" at 800,679 size 78x59; TextOff 'Text'
   Button "Template_Button_3" at 720,679 size 78x59; TextOff 'Text'
   Button "Template_Button_4" at 640,679 size 78x59; TextOff 'Text'
   Button "Template_Button_5" at 561,679 size 78x59; TextOff 'Text'
   Button "Template_Button_6" at 481,679 size 78x59; TextOff 'Text'
   Button "Template_Button_7" at 401,679 size 78x59; TextOff 'Text'
   Button "Template_Button_8" at 321,679 size 78x59; TextOff 'Text'
   Button "Template_Button_9" at 241,679 size 78x59; TextOff 'R-3'
      on Release: ActivateScreen("Rolling Stand 3", 0)
   Button "Template_Button_10" at 161,679 size 78x59; TextOff 'R-2'
      on Release: ActivateScreen("Rolling Stand 2", 0)
   Button "Template_Button_11" at 81,679 size 78x59; TextOn 'R-1'; TextOff 'R-1'
      on Release: ActivateScreen("Rolling Stand 1", 0)
   Button "Start screen" at 1,679 size 78x59; TextOn 'Start screen'; TextOff 'Start screen'; PictureOn "NavigateHome_TP1500_Comfort_TR"; PictureOff "NavigateHome_TP1500_Comfort_TR"
      on Release: ActivateScreen("Home", 0)
   AlarmView "Alarm view_Unacknowledged" at 0,0 size 1280x23
*)